(* Logix 5000 project; controller PLC_MCC1300_75F1 vendor 1 type 14 code 166 rev 32.11; software revision 32.04; part 45 of 83 *)
(* tags used below, declared in another part *)
   CONST_tPlant : UDT_PLANT_CONSTANTS;
   GP_PosWindow : GP_PosWindow;
   GP_TrackingSearchPlate : GP_TrackingSearchPlate;
   GP_TrackingValidateIndex : GP_TrackingValidateIndex;
   M30xTrimDeck : MAC_TrimmingDeck[5];
   M30xTrimDeck_DATA : UDT_ConvoyCap_ZC[5];
   M30xTrimDeck_HMR : MAC_TrimmingDeck_HMR[5];
   M30xTrimDeck_HMW : MAC_TrimmingDeck_HMW[5];
   TMP_d : DINT;
   TMP_dBufferIndex : DINT;
   TMP_dIndex : DINT;
   xAlwaysOFF : BOOL;
   xAlwaysON : BOOL;
   Z300_BufferPlate : UDT_LINE_BUFFER_PLATE;
   Z300_LineTracking : UDT_LINE_TRACKING;
   Z301 : MAC_Zone_ML;
(* MainProgram, continued *)

ROUTINE M30xTrimDeck_Logic   (* ladder *)
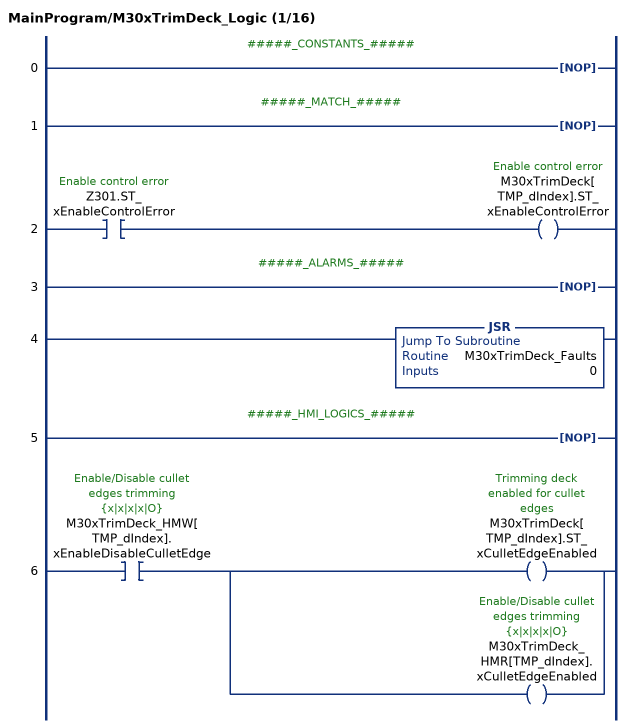
   // #####_CONSTANTS_#####
   0: NOP();
   // #####_MATCH_#####
   1: NOP();
   2: XIC(Z301.ST_xEnableControlError)OTE(M30xTrimDeck[TMP_dIndex].ST_xEnableControlError);
   // #####_ALARMS_#####
   3: NOP();
   4: JSR(M30xTrimDeck_Faults,0);
   // #####_HMI_LOGICS_#####
   5: NOP();
   6: XIC(M30xTrimDeck_HMW[TMP_dIndex].xEnableDisableCulletEdge)[OTE(M30xTrimDeck[TMP_dIndex].ST_xCulletEdgeEnabled) ,OTE(M30xTrimDeck_HMR[TMP_dIndex].xCulletEdgeEnabled) ];
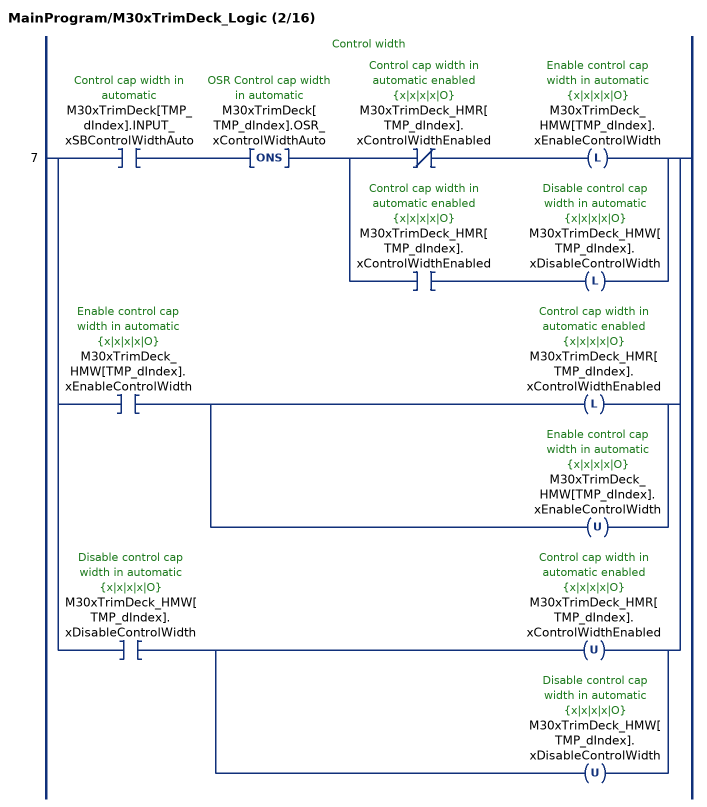
   // Control width
   7: [XIC(M30xTrimDeck[TMP_dIndex].INPUT_xSBControlWidthAuto) ONS(M30xTrimDeck[TMP_dIndex].OSR_xControlWidthAuto) [XIO(M30xTrimDeck_HMR[TMP_dIndex].xControlWidthEnabled) OTL(M30xTrimDeck_HMW[TMP_dIndex].xEnableControlWidth) ,XIC(M30xTrimDeck_HMR[TMP_dIndex].xControlWidthEnabled) OTL(M30xTrimDeck_HMW[TMP_dIndex].xDisableControlWidth) ] ,[XIC(M30xTrimDeck_HMW[TMP_dIndex].xEnableControlWidth) [OTL(M30xTrimDeck_HMR[TMP_dIndex].xControlWidthEnabled) ,OTU(M30xTrimDeck_HMW[TMP_dIndex].xEnableControlWidth) ] ,XIC(M30xTrimDeck_HMW[TMP_dIndex].xDisableControlWidth) [OTU(M30xTrimDeck_HMR[TMP_dIndex].xControlWidthEnabled) ,OTU(M30xTrimDeck_HMW[TMP_dIndex].xDisableControlWidth) ] ] ];
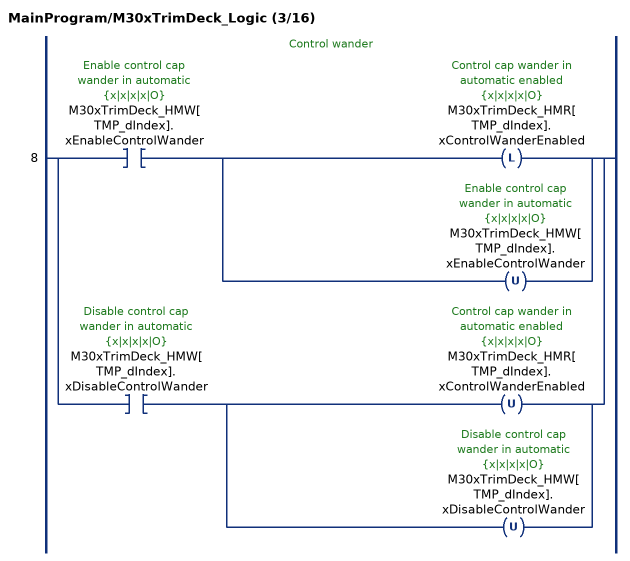
   // Control wander
   8: [XIC(M30xTrimDeck_HMW[TMP_dIndex].xEnableControlWander) [OTL(M30xTrimDeck_HMR[TMP_dIndex].xControlWanderEnabled) ,OTU(M30xTrimDeck_HMW[TMP_dIndex].xEnableControlWander) ] ,XIC(M30xTrimDeck_HMW[TMP_dIndex].xDisableControlWander) [OTU(M30xTrimDeck_HMR[TMP_dIndex].xControlWanderEnabled) ,OTU(M30xTrimDeck_HMW[TMP_dIndex].xDisableControlWander) ] ];
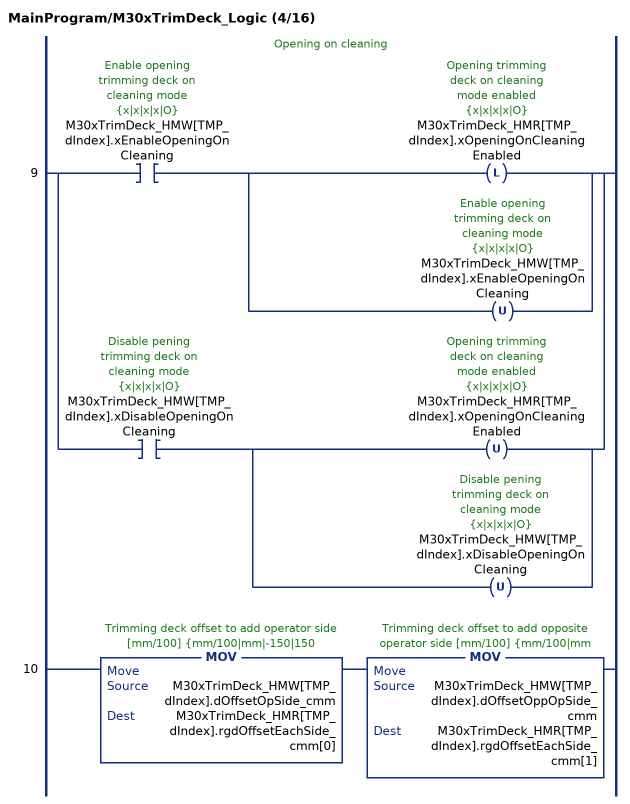
   // Opening on cleaning
   9: [XIC(M30xTrimDeck_HMW[TMP_dIndex].xEnableOpeningOnCleaning) [OTL(M30xTrimDeck_HMR[TMP_dIndex].xOpeningOnCleaningEnabled) ,OTU(M30xTrimDeck_HMW[TMP_dIndex].xEnableOpeningOnCleaning) ] ,XIC(M30xTrimDeck_HMW[TMP_dIndex].xDisableOpeningOnCleaning) [OTU(M30xTrimDeck_HMR[TMP_dIndex].xOpeningOnCleaningEnabled) ,OTU(M30xTrimDeck_HMW[TMP_dIndex].xDisableOpeningOnCleaning) ] ];
   10: MOV(M30xTrimDeck_HMW[TMP_dIndex].dOffsetOpSide_cmm,M30xTrimDeck_HMR[TMP_dIndex].rgdOffsetEachSide_cmm[0])MOV(M30xTrimDeck_HMW[TMP_dIndex].dOffsetOppOpSide_cmm,M30xTrimDeck_HMR[TMP_dIndex].rgdOffsetEachSide_cmm[1]);
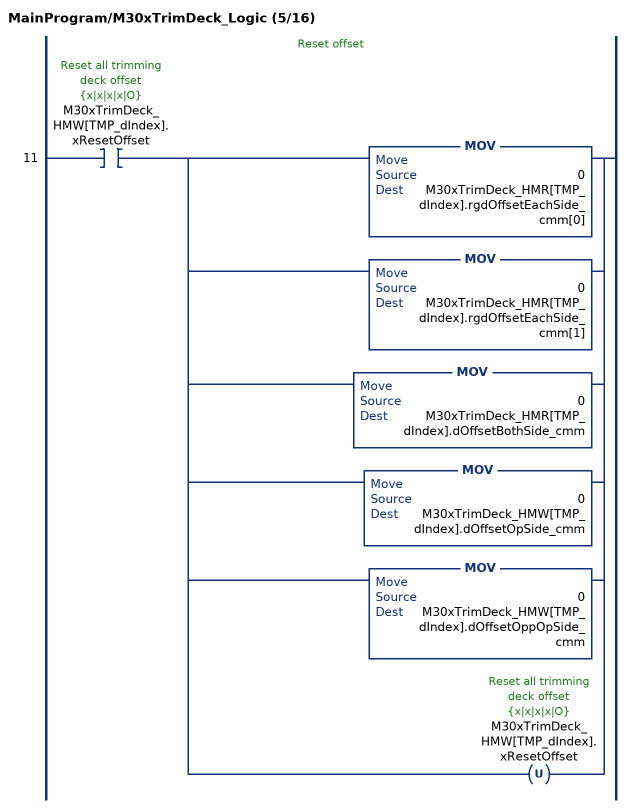
   // Reset offset
   11: XIC(M30xTrimDeck_HMW[TMP_dIndex].xResetOffset)[MOV(0,M30xTrimDeck_HMR[TMP_dIndex].rgdOffsetEachSide_cmm[0]) ,MOV(0,M30xTrimDeck_HMR[TMP_dIndex].rgdOffsetEachSide_cmm[1]) ,MOV(0,M30xTrimDeck_HMR[TMP_dIndex].dOffsetBothSide_cmm) ,MOV(0,M30xTrimDeck_HMW[TMP_dIndex].dOffsetOpSide_cmm) ,MOV(0,M30xTrimDeck_HMW[TMP_dIndex].dOffsetOppOpSide_cmm) ,OTU(M30xTrimDeck_HMW[TMP_dIndex].xResetOffset) ];
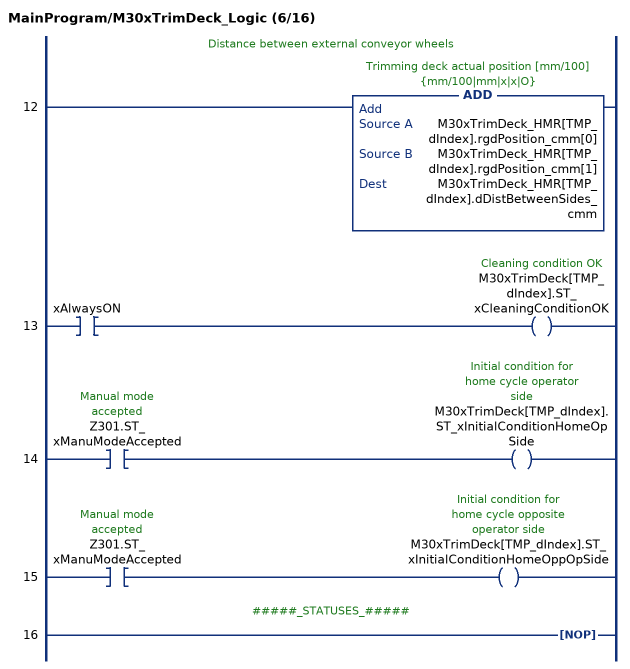
   // Distance between external conveyor wheels
   12: ADD(M30xTrimDeck_HMR[TMP_dIndex].rgdPosition_cmm[0],M30xTrimDeck_HMR[TMP_dIndex].rgdPosition_cmm[1],M30xTrimDeck_HMR[TMP_dIndex].dDistBetweenSides_cmm);
   13: XIC(xAlwaysON)OTE(M30xTrimDeck[TMP_dIndex].ST_xCleaningConditionOK);
   14: XIC(Z301.ST_xManuModeAccepted)OTE(M30xTrimDeck[TMP_dIndex].ST_xInitialConditionHomeOpSide);
   15: XIC(Z301.ST_xManuModeAccepted)OTE(M30xTrimDeck[TMP_dIndex].ST_xInitialConditionHomeOppOpSide);
   // #####_STATUSES_#####
   16: NOP();
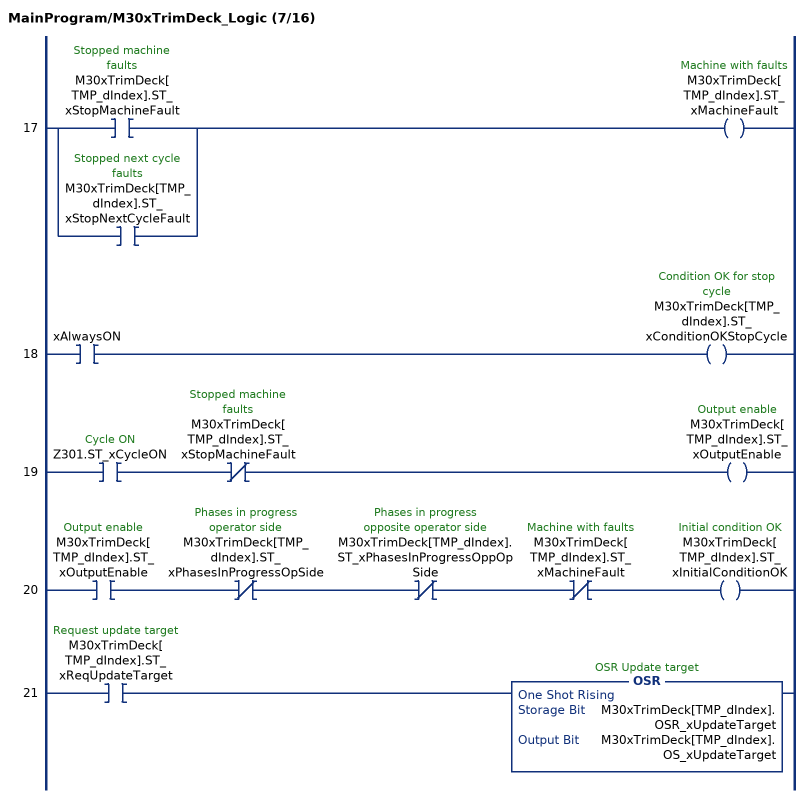
   17: [XIC(M30xTrimDeck[TMP_dIndex].ST_xStopMachineFault) ,XIC(M30xTrimDeck[TMP_dIndex].ST_xStopNextCycleFault) ]OTE(M30xTrimDeck[TMP_dIndex].ST_xMachineFault);
   18: XIC(xAlwaysON)OTE(M30xTrimDeck[TMP_dIndex].ST_xConditionOKStopCycle);
   19: XIC(Z301.ST_xCycleON)XIO(M30xTrimDeck[TMP_dIndex].ST_xStopMachineFault)OTE(M30xTrimDeck[TMP_dIndex].ST_xOutputEnable);
   20: XIC(M30xTrimDeck[TMP_dIndex].ST_xOutputEnable)XIO(M30xTrimDeck[TMP_dIndex].ST_xPhasesInProgressOpSide)XIO(M30xTrimDeck[TMP_dIndex].ST_xPhasesInProgressOppOpSide)XIO(M30xTrimDeck[TMP_dIndex].ST_xMachineFault)OTE(M30xTrimDeck[TMP_dIndex].ST_xInitialConditionOK);
   21: XIC(M30xTrimDeck[TMP_dIndex].ST_xReqUpdateTarget)OSR(M30xTrimDeck[TMP_dIndex].OSR_xUpdateTarget,M30xTrimDeck[TMP_dIndex].OS_xUpdateTarget);
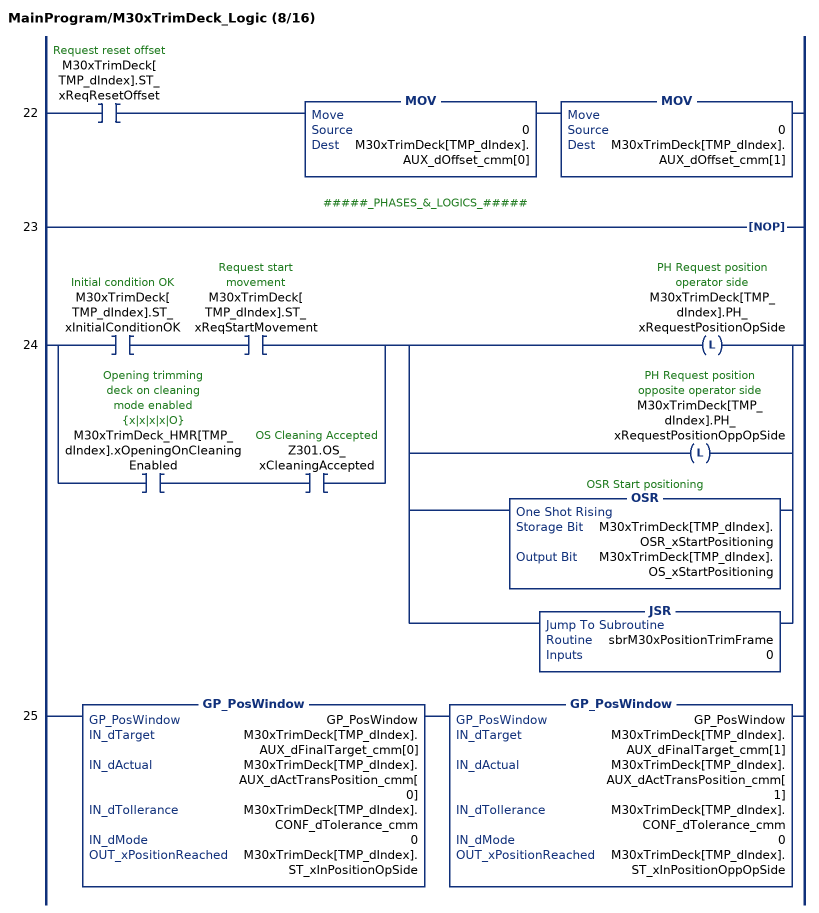
   22: XIC(M30xTrimDeck[TMP_dIndex].ST_xReqResetOffset)MOV(0,M30xTrimDeck[TMP_dIndex].AUX_dOffset_cmm[0])MOV(0,M30xTrimDeck[TMP_dIndex].AUX_dOffset_cmm[1]);
   // #####_PHASES_&_LOGICS_#####
   23: NOP();
   24: [XIC(M30xTrimDeck[TMP_dIndex].ST_xInitialConditionOK) XIC(M30xTrimDeck[TMP_dIndex].ST_xReqStartMovement) ,XIC(M30xTrimDeck_HMR[TMP_dIndex].xOpeningOnCleaningEnabled) XIC(Z301.OS_xCleaningAccepted) ][OTL(M30xTrimDeck[TMP_dIndex].PH_xRequestPositionOpSide) ,OTL(M30xTrimDeck[TMP_dIndex].PH_xRequestPositionOppOpSide) ,OSR(M30xTrimDeck[TMP_dIndex].OSR_xStartPositioning,M30xTrimDeck[TMP_dIndex].OS_xStartPositioning) ,JSR(sbrM30xPositionTrimFrame,0) ];
   25: GP_PosWindow(GP_PosWindow,M30xTrimDeck[TMP_dIndex].AUX_dFinalTarget_cmm[0],M30xTrimDeck[TMP_dIndex].AUX_dActTransPosition_cmm[0],M30xTrimDeck[TMP_dIndex].CONF_dTolerance_cmm,0,M30xTrimDeck[TMP_dIndex].ST_xInPositionOpSide)GP_PosWindow(GP_PosWindow,M30xTrimDeck[TMP_dIndex].AUX_dFinalTarget_cmm[1],M30xTrimDeck[TMP_dIndex].AUX_dActTransPosition_cmm[1],M30xTrimDeck[TMP_dIndex].CONF_dTolerance_cmm,0,M30xTrimDeck[TMP_dIndex].ST_xInPositionOppOpSide);
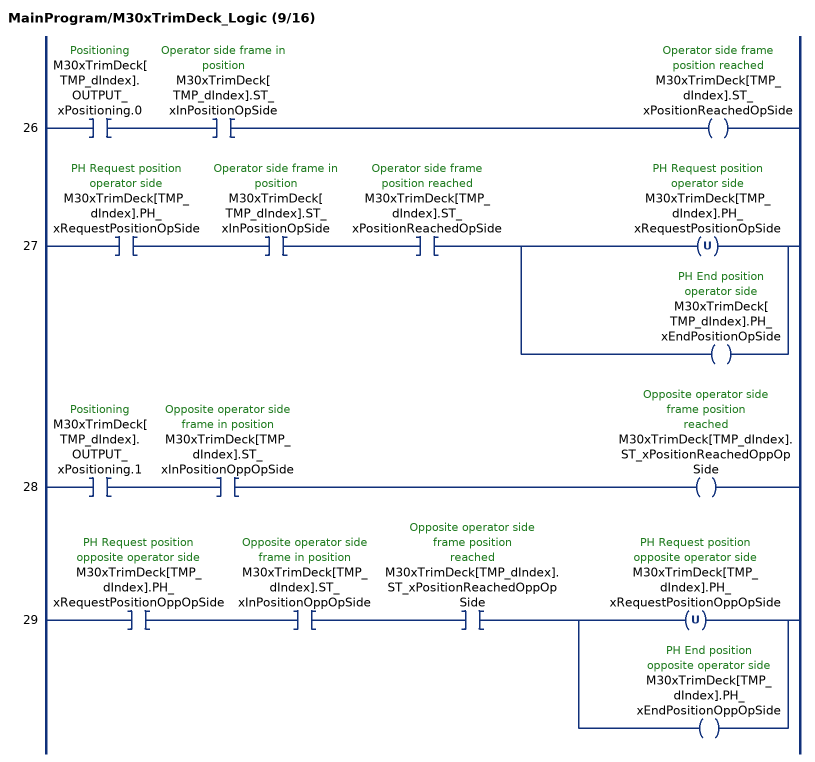
   26: XIC(M30xTrimDeck[TMP_dIndex].OUTPUT_xPositioning.0)XIC(M30xTrimDeck[TMP_dIndex].ST_xInPositionOpSide)OTE(M30xTrimDeck[TMP_dIndex].ST_xPositionReachedOpSide);
   27: XIC(M30xTrimDeck[TMP_dIndex].PH_xRequestPositionOpSide)XIC(M30xTrimDeck[TMP_dIndex].ST_xInPositionOpSide)XIC(M30xTrimDeck[TMP_dIndex].ST_xPositionReachedOpSide)[OTU(M30xTrimDeck[TMP_dIndex].PH_xRequestPositionOpSide) ,OTE(M30xTrimDeck[TMP_dIndex].PH_xEndPositionOpSide) ];
   28: XIC(M30xTrimDeck[TMP_dIndex].OUTPUT_xPositioning.1)XIC(M30xTrimDeck[TMP_dIndex].ST_xInPositionOppOpSide)OTE(M30xTrimDeck[TMP_dIndex].ST_xPositionReachedOppOpSide);
   29: XIC(M30xTrimDeck[TMP_dIndex].PH_xRequestPositionOppOpSide)XIC(M30xTrimDeck[TMP_dIndex].ST_xInPositionOppOpSide)XIC(M30xTrimDeck[TMP_dIndex].ST_xPositionReachedOppOpSide)[OTU(M30xTrimDeck[TMP_dIndex].PH_xRequestPositionOppOpSide) ,OTE(M30xTrimDeck[TMP_dIndex].PH_xEndPositionOppOpSide) ];
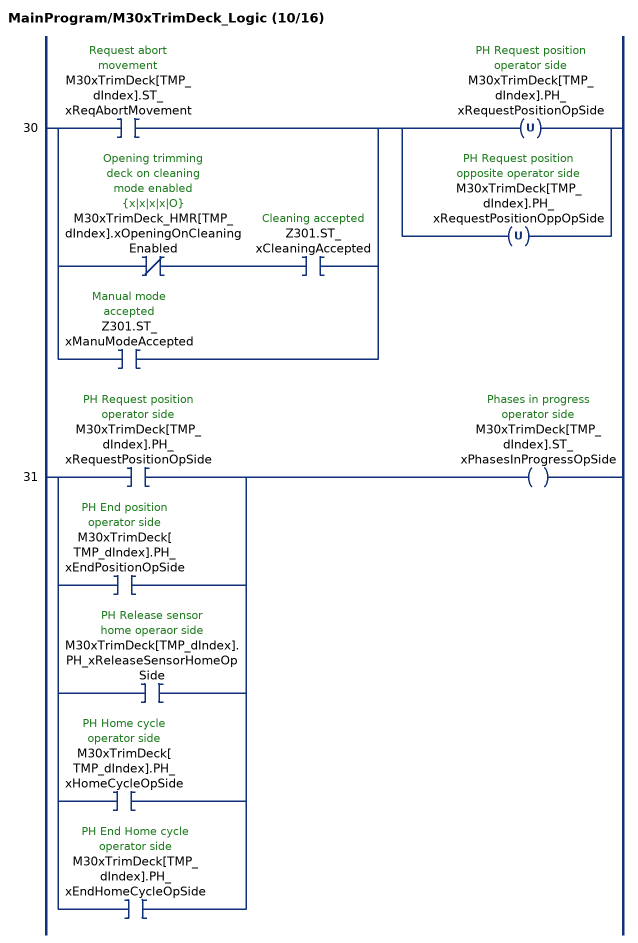
   30: [XIC(M30xTrimDeck[TMP_dIndex].ST_xReqAbortMovement) ,XIO(M30xTrimDeck_HMR[TMP_dIndex].xOpeningOnCleaningEnabled) XIC(Z301.ST_xCleaningAccepted) ,XIC(Z301.ST_xManuModeAccepted) ][OTU(M30xTrimDeck[TMP_dIndex].PH_xRequestPositionOpSide) ,OTU(M30xTrimDeck[TMP_dIndex].PH_xRequestPositionOppOpSide) ];
   31: [XIC(M30xTrimDeck[TMP_dIndex].PH_xRequestPositionOpSide) ,XIC(M30xTrimDeck[TMP_dIndex].PH_xEndPositionOpSide) ,XIC(M30xTrimDeck[TMP_dIndex].PH_xReleaseSensorHomeOpSide) ,XIC(M30xTrimDeck[TMP_dIndex].PH_xHomeCycleOpSide) ,XIC(M30xTrimDeck[TMP_dIndex].PH_xEndHomeCycleOpSide) ]OTE(M30xTrimDeck[TMP_dIndex].ST_xPhasesInProgressOpSide);
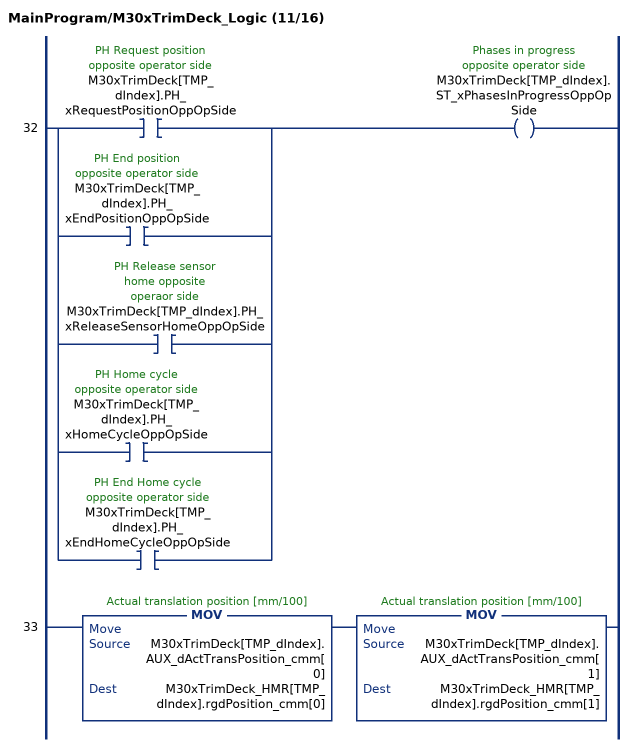
   32: [XIC(M30xTrimDeck[TMP_dIndex].PH_xRequestPositionOppOpSide) ,XIC(M30xTrimDeck[TMP_dIndex].PH_xEndPositionOppOpSide) ,XIC(M30xTrimDeck[TMP_dIndex].PH_xReleaseSensorHomeOppOpSide) ,XIC(M30xTrimDeck[TMP_dIndex].PH_xHomeCycleOppOpSide) ,XIC(M30xTrimDeck[TMP_dIndex].PH_xEndHomeCycleOppOpSide) ]OTE(M30xTrimDeck[TMP_dIndex].ST_xPhasesInProgressOppOpSide);
   33: MOV(M30xTrimDeck[TMP_dIndex].AUX_dActTransPosition_cmm[0],M30xTrimDeck_HMR[TMP_dIndex].rgdPosition_cmm[0])MOV(M30xTrimDeck[TMP_dIndex].AUX_dActTransPosition_cmm[1],M30xTrimDeck_HMR[TMP_dIndex].rgdPosition_cmm[1]);
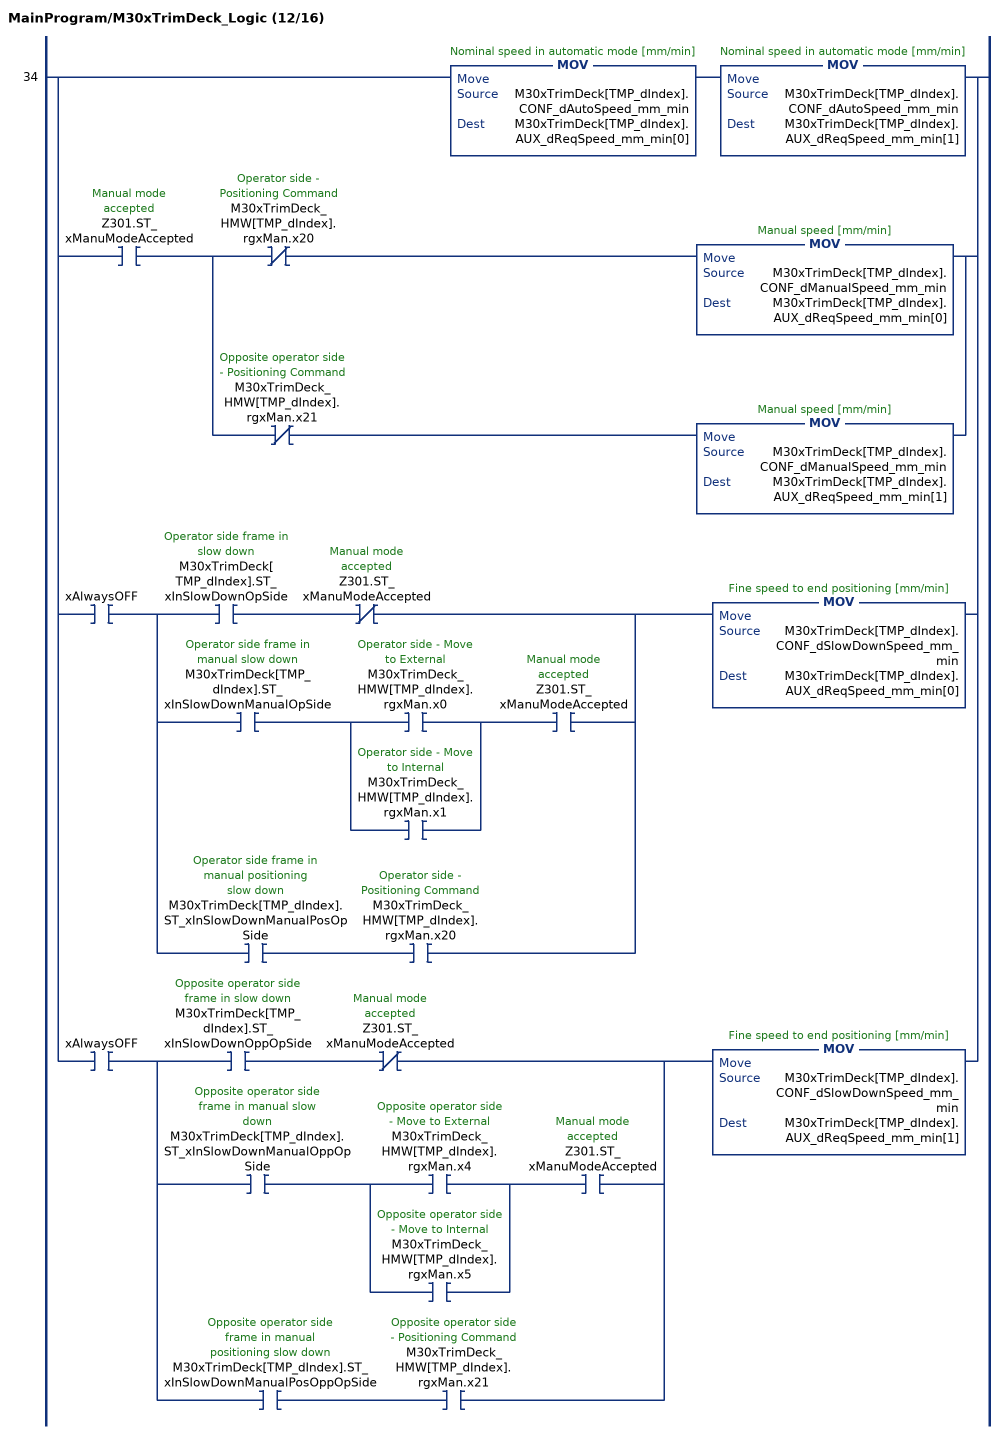
   34: [MOV(M30xTrimDeck[TMP_dIndex].CONF_dAutoSpeed_mm_min,M30xTrimDeck[TMP_dIndex].AUX_dReqSpeed_mm_min[0]) MOV(M30xTrimDeck[TMP_dIndex].CONF_dAutoSpeed_mm_min,M30xTrimDeck[TMP_dIndex].AUX_dReqSpeed_mm_min[1]) ,XIC(Z301.ST_xManuModeAccepted) [XIO(M30xTrimDeck_HMW[TMP_dIndex].rgxMan.x20) MOV(M30xTrimDeck[TMP_dIndex].CONF_dManualSpeed_mm_min,M30xTrimDeck[TMP_dIndex].AUX_dReqSpeed_mm_min[0]) ,XIO(M30xTrimDeck_HMW[TMP_dIndex].rgxMan.x21) MOV(M30xTrimDeck[TMP_dIndex].CONF_dManualSpeed_mm_min,M30xTrimDeck[TMP_dIndex].AUX_dReqSpeed_mm_min[1]) ] ,XIC(xAlwaysOFF) [XIC(M30xTrimDeck[TMP_dIndex].ST_xInSlowDownOpSide) XIO(Z301.ST_xManuModeAccepted) ,XIC(M30xTrimDeck[TMP_dIndex].ST_xInSlowDownManualOpSide) [XIC(M30xTrimDeck_HMW[TMP_dIndex].rgxMan.x0) ,XIC(M30xTrimDeck_HMW[TMP_dIndex].rgxMan.x1) ] XIC(Z301.ST_xManuModeAccepted) ,XIC(M30xTrimDeck[TMP_dIndex].ST_xInSlowDownManualPosOpSide) XIC(M30xTrimDeck_HMW[TMP_dIndex].rgxMan.x20) ] MOV(M30xTrimDeck[TMP_dIndex].CONF_dSlowDownSpeed_mm_min,M30xTrimDeck[TMP_dIndex].AUX_dReqSpeed_mm_min[0]) ,XIC(xAlwaysOFF) [XIC(M30xTrimDeck[TMP_dIndex].ST_xInSlowDownOppOpSide) XIO(Z301.ST_xManuModeAccepted) ,XIC(M30xTrimDeck[TMP_dIndex].ST_xInSlowDownManualOppOpSide) [XIC(M30xTrimDeck_HMW[TMP_dIndex].rgxMan.x4) ,XIC(M30xTrimDeck_HMW[TMP_dIndex].rgxMan.x5) ] XIC(Z301.ST_xManuModeAccepted) ,XIC(M30xTrimDeck[TMP_dIndex].ST_xInSlowDownManualPosOppOpSide) XIC(M30xTrimDeck_HMW[TMP_dIndex].rgxMan.x21) ] MOV(M30xTrimDeck[TMP_dIndex].CONF_dSlowDownSpeed_mm_min,M30xTrimDeck[TMP_dIndex].AUX_dReqSpeed_mm_min[1]) ];